REGION Network 28
   #temp := SCALE(IN := "5#净环热水阀门开度",
                  HI_LIM := 100.0,
                  LO_LIM := 0.0,
                  BIPOLAR := "AlwaysFALSE",
                  OUT => "AI"."5#净环热水阀门开度");
END_REGION

REGION Network 29
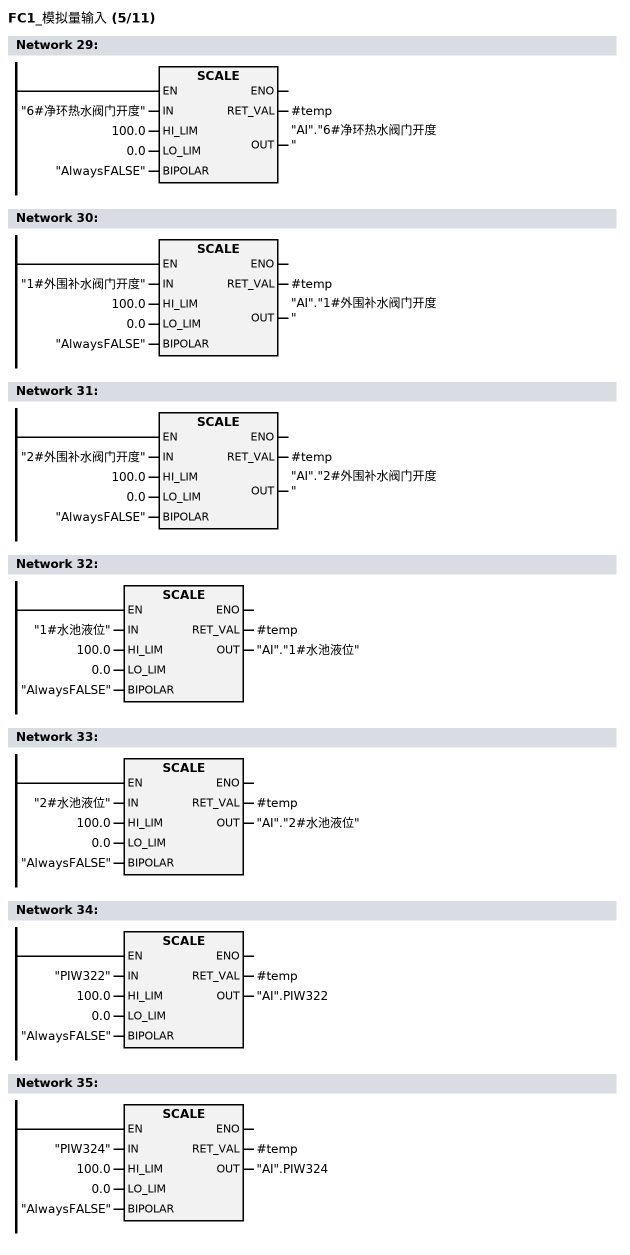
   #temp := SCALE(IN := "6#净环热水阀门开度",
                  HI_LIM := 100.0,
                  LO_LIM := 0.0,
                  BIPOLAR := "AlwaysFALSE",
                  OUT => "AI"."6#净环热水阀门开度");
END_REGION

REGION Network 30
   #temp := SCALE(IN := "1#外围补水阀门开度",
                  HI_LIM := 100.0,
                  LO_LIM := 0.0,
                  BIPOLAR := "AlwaysFALSE",
                  OUT => "AI"."1#外围补水阀门开度");
END_REGION

REGION Network 31
   #temp := SCALE(IN := "2#外围补水阀门开度",
                  HI_LIM := 100.0,
                  LO_LIM := 0.0,
                  BIPOLAR := "AlwaysFALSE",
                  OUT => "AI"."2#外围补水阀门开度");
END_REGION

REGION Network 32
   #temp := SCALE(IN := "1#水池液位",
                  HI_LIM := 100.0,
                  LO_LIM := 0.0,
                  BIPOLAR := "AlwaysFALSE",
                  OUT => "AI"."1#水池液位");
END_REGION

REGION Network 33
   #temp := SCALE(IN := "2#水池液位",
                  HI_LIM := 100.0,
                  LO_LIM := 0.0,
                  BIPOLAR := "AlwaysFALSE",
                  OUT => "AI"."2#水池液位");
END_REGION

REGION Network 34
   #temp := SCALE(IN := "PIW322", HI_LIM := 100.0, LO_LIM := 0.0, BIPOLAR := "AlwaysFALSE", OUT => "AI".PIW322);
END_REGION

REGION Network 35
   #temp := SCALE(IN := "PIW324", HI_LIM := 100.0, LO_LIM := 0.0, BIPOLAR := "AlwaysFALSE", OUT => "AI".PIW324);
END_REGION

REGION Network 36
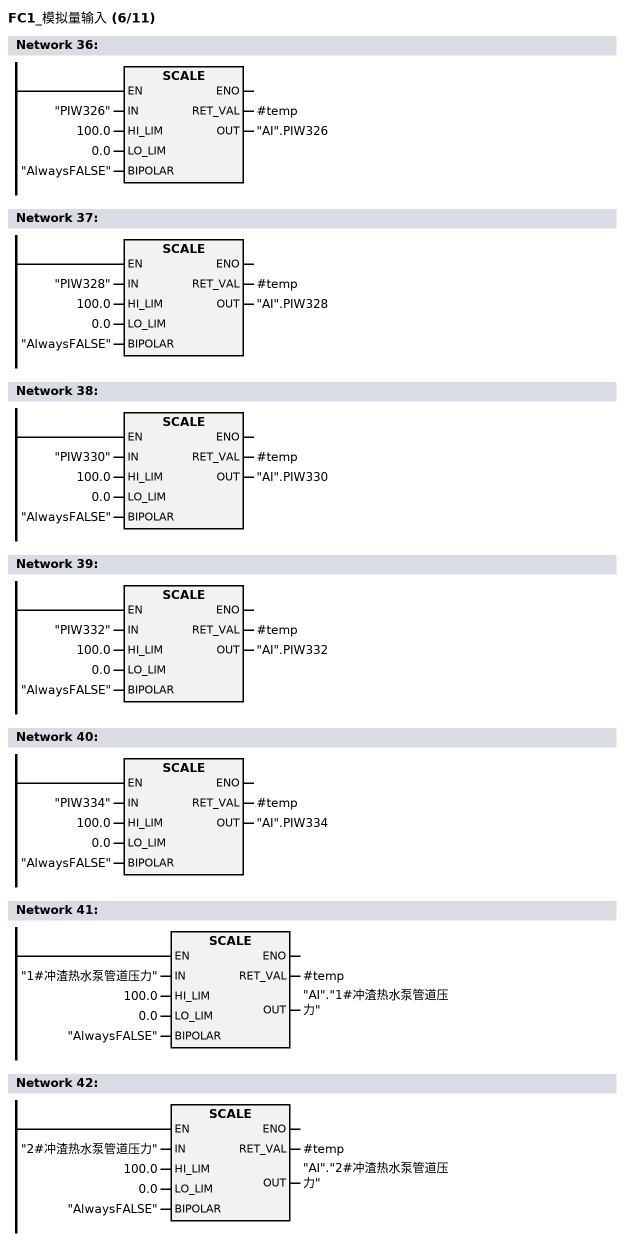
   #temp := SCALE(IN := "PIW326", HI_LIM := 100.0, LO_LIM := 0.0, BIPOLAR := "AlwaysFALSE", OUT => "AI".PIW326);
END_REGION

REGION Network 37
   #temp := SCALE(IN := "PIW328", HI_LIM := 100.0, LO_LIM := 0.0, BIPOLAR := "AlwaysFALSE", OUT => "AI".PIW328);
END_REGION

REGION Network 38
   #temp := SCALE(IN := "PIW330", HI_LIM := 100.0, LO_LIM := 0.0, BIPOLAR := "AlwaysFALSE", OUT => "AI".PIW330);
END_REGION

REGION Network 39
   #temp := SCALE(IN := "PIW332", HI_LIM := 100.0, LO_LIM := 0.0, BIPOLAR := "AlwaysFALSE", OUT => "AI".PIW332);
END_REGION

REGION Network 40
   #temp := SCALE(IN := "PIW334", HI_LIM := 100.0, LO_LIM := 0.0, BIPOLAR := "AlwaysFALSE", OUT => "AI".PIW334);
END_REGION

REGION Network 41
   #temp := SCALE(IN := "1#冲渣热水泵管道压力",
                  HI_LIM := 100.0,
                  LO_LIM := 0.0,
                  BIPOLAR := "AlwaysFALSE",
                  OUT => "AI"."1#冲渣热水泵管道压力");
END_REGION

REGION Network 42
   #temp := SCALE(IN := "2#冲渣热水泵管道压力",
                  HI_LIM := 100.0,
                  LO_LIM := 0.0,
                  BIPOLAR := "AlwaysFALSE",
                  OUT => "AI"."2#冲渣热水泵管道压力");
END_REGION

REGION Network 43
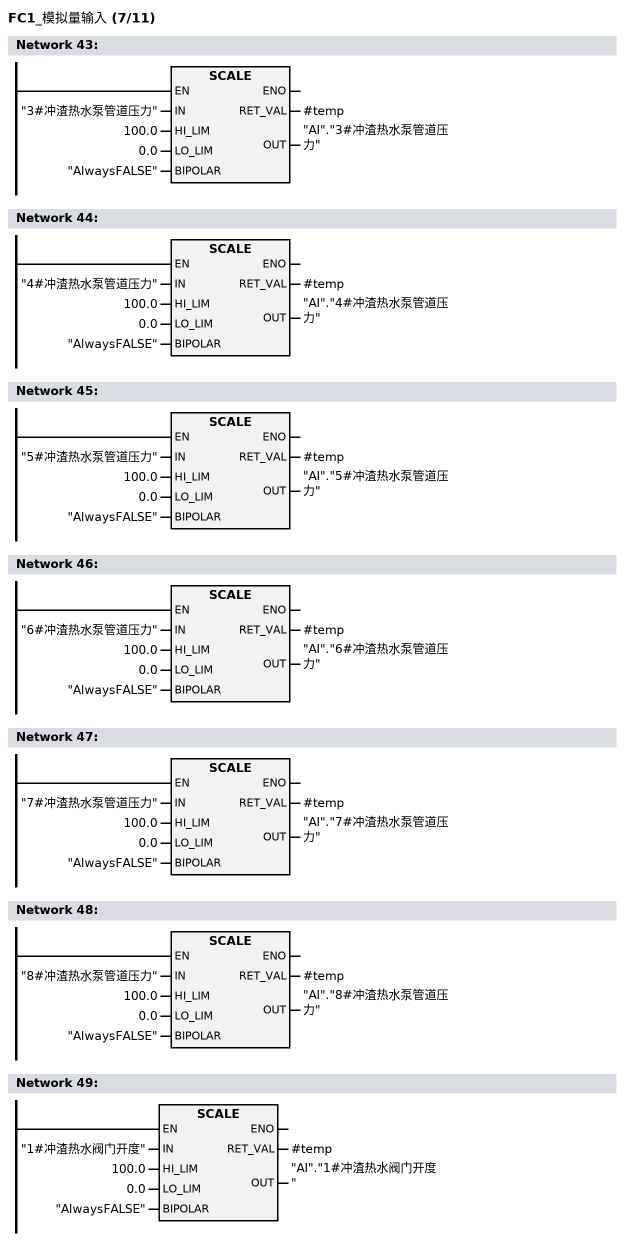
   #temp := SCALE(IN := "3#冲渣热水泵管道压力",
                  HI_LIM := 100.0,
                  LO_LIM := 0.0,
                  BIPOLAR := "AlwaysFALSE",
                  OUT => "AI"."3#冲渣热水泵管道压力");
END_REGION

REGION Network 44
   #temp := SCALE(IN := "4#冲渣热水泵管道压力",
                  HI_LIM := 100.0,
                  LO_LIM := 0.0,
                  BIPOLAR := "AlwaysFALSE",
                  OUT => "AI"."4#冲渣热水泵管道压力");
END_REGION

REGION Network 45
   #temp := SCALE(IN := "5#冲渣热水泵管道压力",
                  HI_LIM := 100.0,
                  LO_LIM := 0.0,
                  BIPOLAR := "AlwaysFALSE",
                  OUT => "AI"."5#冲渣热水泵管道压力");
END_REGION

REGION Network 46
   #temp := SCALE(IN := "6#冲渣热水泵管道压力",
                  HI_LIM := 100.0,
                  LO_LIM := 0.0,
                  BIPOLAR := "AlwaysFALSE",
                  OUT => "AI"."6#冲渣热水泵管道压力");
END_REGION

REGION Network 47
   #temp := SCALE(IN := "7#冲渣热水泵管道压力",
                  HI_LIM := 100.0,
                  LO_LIM := 0.0,
                  BIPOLAR := "AlwaysFALSE",
                  OUT => "AI"."7#冲渣热水泵管道压力");
END_REGION

REGION Network 48
   #temp := SCALE(IN := "8#冲渣热水泵管道压力",
                  HI_LIM := 100.0,
                  LO_LIM := 0.0,
                  BIPOLAR := "AlwaysFALSE",
                  OUT => "AI"."8#冲渣热水泵管道压力");
END_REGION

REGION Network 49
   #temp := SCALE(IN := "1#冲渣热水阀门开度",
                  HI_LIM := 100.0,
                  LO_LIM := 0.0,
                  BIPOLAR := "AlwaysFALSE",
                  OUT => "AI"."1#冲渣热水阀门开度");
END_REGION

REGION Network 50
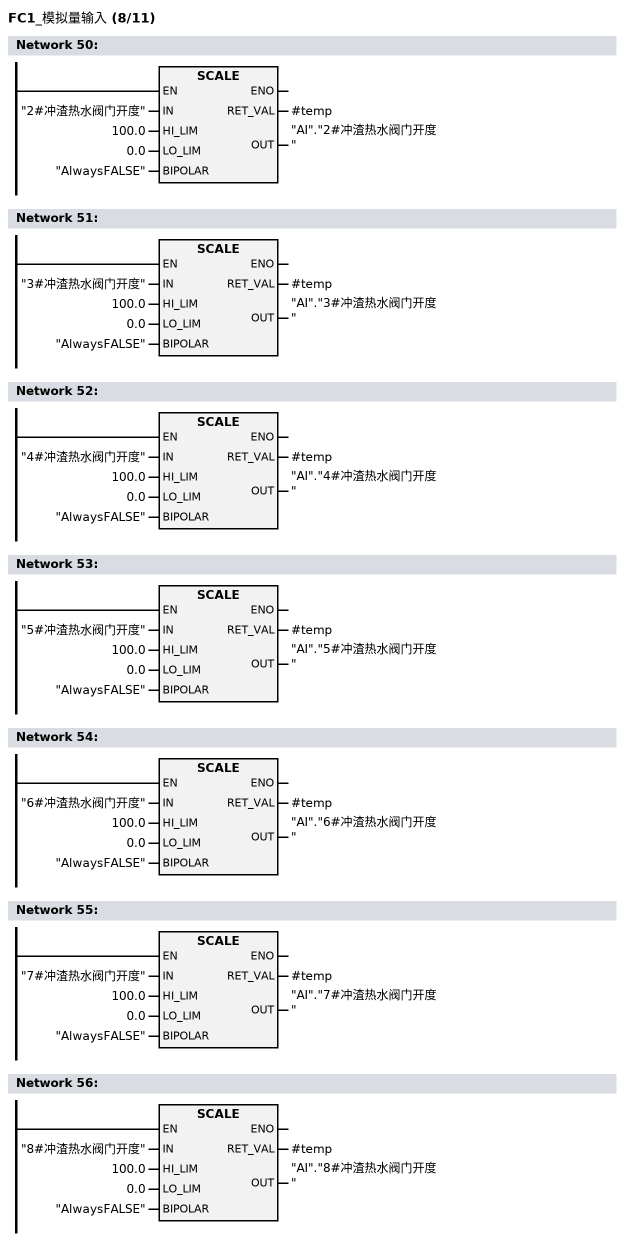
   #temp := SCALE(IN := "2#冲渣热水阀门开度",
                  HI_LIM := 100.0,
                  LO_LIM := 0.0,
                  BIPOLAR := "AlwaysFALSE",
                  OUT => "AI"."2#冲渣热水阀门开度");
END_REGION

REGION Network 51
   #temp := SCALE(IN := "3#冲渣热水阀门开度",
                  HI_LIM := 100.0,
                  LO_LIM := 0.0,
                  BIPOLAR := "AlwaysFALSE",
                  OUT => "AI"."3#冲渣热水阀门开度");
END_REGION

REGION Network 52
   #temp := SCALE(IN := "4#冲渣热水阀门开度",
                  HI_LIM := 100.0,
                  LO_LIM := 0.0,
                  BIPOLAR := "AlwaysFALSE",
                  OUT => "AI"."4#冲渣热水阀门开度");
END_REGION

REGION Network 53
   #temp := SCALE(IN := "5#冲渣热水阀门开度",
                  HI_LIM := 100.0,
                  LO_LIM := 0.0,
                  BIPOLAR := "AlwaysFALSE",
                  OUT => "AI"."5#冲渣热水阀门开度");
END_REGION

REGION Network 54
   #temp := SCALE(IN := "6#冲渣热水阀门开度",
                  HI_LIM := 100.0,
                  LO_LIM := 0.0,
                  BIPOLAR := "AlwaysFALSE",
                  OUT => "AI"."6#冲渣热水阀门开度");
END_REGION

REGION Network 55
   #temp := SCALE(IN := "7#冲渣热水阀门开度",
                  HI_LIM := 100.0,
                  LO_LIM := 0.0,
                  BIPOLAR := "AlwaysFALSE",
                  OUT => "AI"."7#冲渣热水阀门开度");
END_REGION

REGION Network 56
   #temp := SCALE(IN := "8#冲渣热水阀门开度",
                  HI_LIM := 100.0,
                  LO_LIM := 0.0,
                  BIPOLAR := "AlwaysFALSE",
                  OUT => "AI"."8#冲渣热水阀门开度");
END_REGION

REGION Network 57
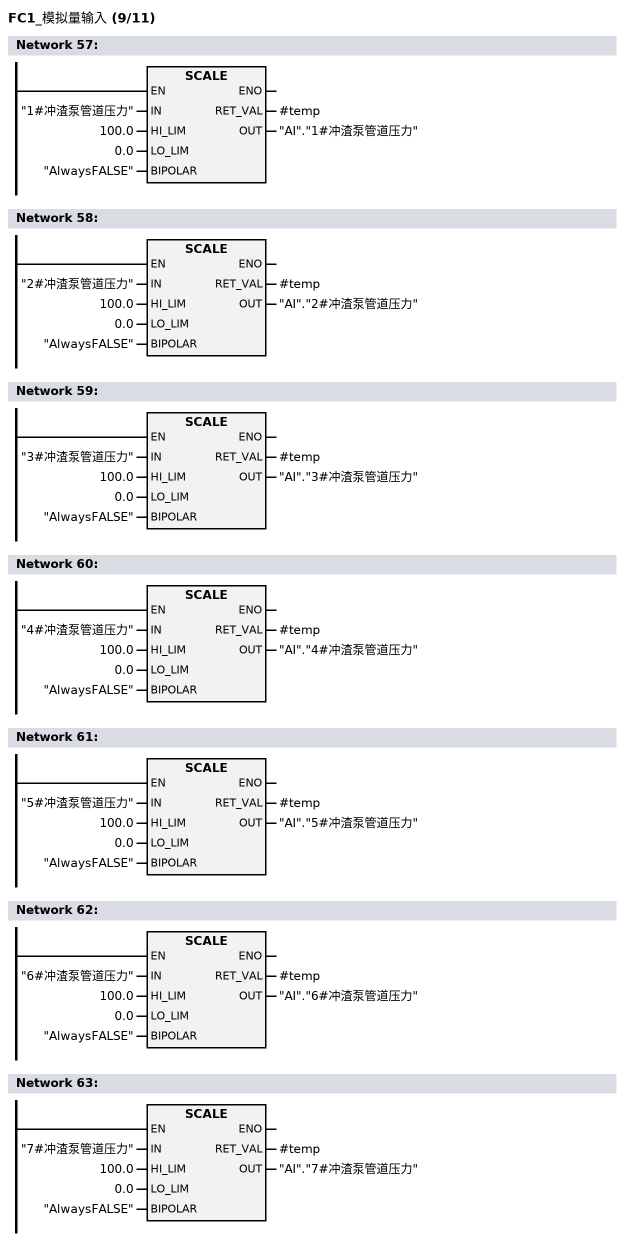
   #temp := SCALE(IN := "1#冲渣泵管道压力",
                  HI_LIM := 100.0,
                  LO_LIM := 0.0,
                  BIPOLAR := "AlwaysFALSE",
                  OUT => "AI"."1#冲渣泵管道压力");
END_REGION

REGION Network 58
   #temp := SCALE(IN := "2#冲渣泵管道压力",
                  HI_LIM := 100.0,
                  LO_LIM := 0.0,
                  BIPOLAR := "AlwaysFALSE",
                  OUT => "AI"."2#冲渣泵管道压力");
END_REGION

REGION Network 59
   #temp := SCALE(IN := "3#冲渣泵管道压力",
                  HI_LIM := 100.0,
                  LO_LIM := 0.0,
                  BIPOLAR := "AlwaysFALSE",
                  OUT => "AI"."3#冲渣泵管道压力");
END_REGION

REGION Network 60
   #temp := SCALE(IN := "4#冲渣泵管道压力",
                  HI_LIM := 100.0,
                  LO_LIM := 0.0,
                  BIPOLAR := "AlwaysFALSE",
                  OUT => "AI"."4#冲渣泵管道压力");
END_REGION

REGION Network 61
   #temp := SCALE(IN := "5#冲渣泵管道压力",
                  HI_LIM := 100.0,
                  LO_LIM := 0.0,
                  BIPOLAR := "AlwaysFALSE",
                  OUT => "AI"."5#冲渣泵管道压力");
END_REGION

REGION Network 62
   #temp := SCALE(IN := "6#冲渣泵管道压力",
                  HI_LIM := 100.0,
                  LO_LIM := 0.0,
                  BIPOLAR := "AlwaysFALSE",
                  OUT => "AI"."6#冲渣泵管道压力");
END_REGION

REGION Network 63
   #temp := SCALE(IN := "7#冲渣泵管道压力",
                  HI_LIM := 100.0,
                  LO_LIM := 0.0,
                  BIPOLAR := "AlwaysFALSE",
                  OUT => "AI"."7#冲渣泵管道压力");
END_REGION

REGION Network 64
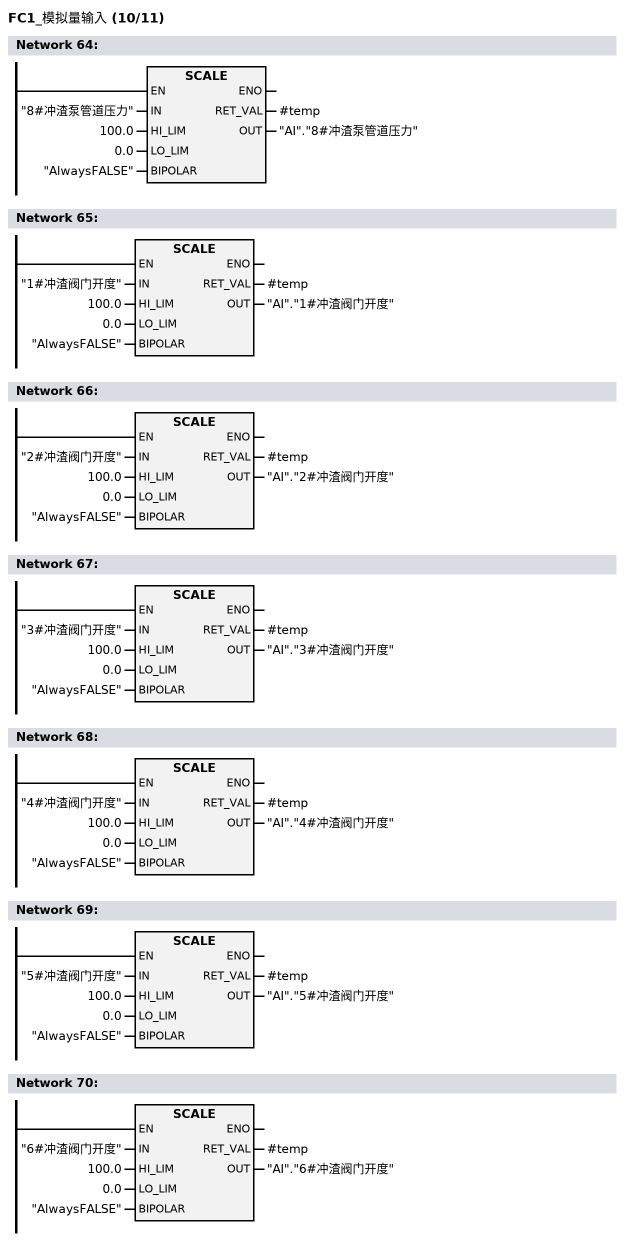
   #temp := SCALE(IN := "8#冲渣泵管道压力",
                  HI_LIM := 100.0,
                  LO_LIM := 0.0,
                  BIPOLAR := "AlwaysFALSE",
                  OUT => "AI"."8#冲渣泵管道压力");
END_REGION

REGION Network 65
   #temp := SCALE(IN := "1#冲渣阀门开度",
                  HI_LIM := 100.0,
                  LO_LIM := 0.0,
                  BIPOLAR := "AlwaysFALSE",
                  OUT => "AI"."1#冲渣阀门开度");
END_REGION

REGION Network 66
   #temp := SCALE(IN := "2#冲渣阀门开度",
                  HI_LIM := 100.0,
                  LO_LIM := 0.0,
                  BIPOLAR := "AlwaysFALSE",
                  OUT => "AI"."2#冲渣阀门开度");
END_REGION

REGION Network 67
   #temp := SCALE(IN := "3#冲渣阀门开度",
                  HI_LIM := 100.0,
                  LO_LIM := 0.0,
                  BIPOLAR := "AlwaysFALSE",
                  OUT => "AI"."3#冲渣阀门开度");
END_REGION

REGION Network 68
   #temp := SCALE(IN := "4#冲渣阀门开度",
                  HI_LIM := 100.0,
                  LO_LIM := 0.0,
                  BIPOLAR := "AlwaysFALSE",
                  OUT => "AI"."4#冲渣阀门开度");
END_REGION

REGION Network 69
   #temp := SCALE(IN := "5#冲渣阀门开度",
                  HI_LIM := 100.0,
                  LO_LIM := 0.0,
                  BIPOLAR := "AlwaysFALSE",
                  OUT => "AI"."5#冲渣阀门开度");
END_REGION

REGION Network 70
   #temp := SCALE(IN := "6#冲渣阀门开度",
                  HI_LIM := 100.0,
                  LO_LIM := 0.0,
                  BIPOLAR := "AlwaysFALSE",
                  OUT => "AI"."6#冲渣阀门开度");
END_REGION

REGION Network 71
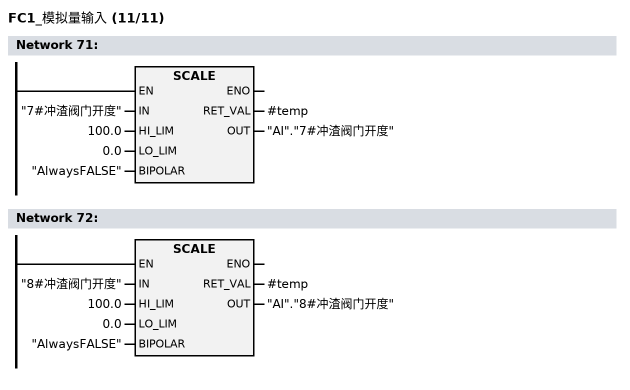
   #temp := SCALE(IN := "7#冲渣阀门开度",
                  HI_LIM := 100.0,
                  LO_LIM := 0.0,
                  BIPOLAR := "AlwaysFALSE",
                  OUT => "AI"."7#冲渣阀门开度");
END_REGION

REGION Network 72
   #temp := SCALE(IN := "8#冲渣阀门开度",
                  HI_LIM := 100.0,
                  LO_LIM := 0.0,
                  BIPOLAR := "AlwaysFALSE",
                  OUT => "AI"."8#冲渣阀门开度");
END_REGION
END_FUNCTION

FUNCTION "FC2_模拟量输出" : Void   // FC2, LAD
{ S7_Optimized_Access := 'TRUE' }
VERSION : 0.1
   VAR_TEMP
      temp_AO : Word;
   END_VAR
BEGIN

REGION Network 1
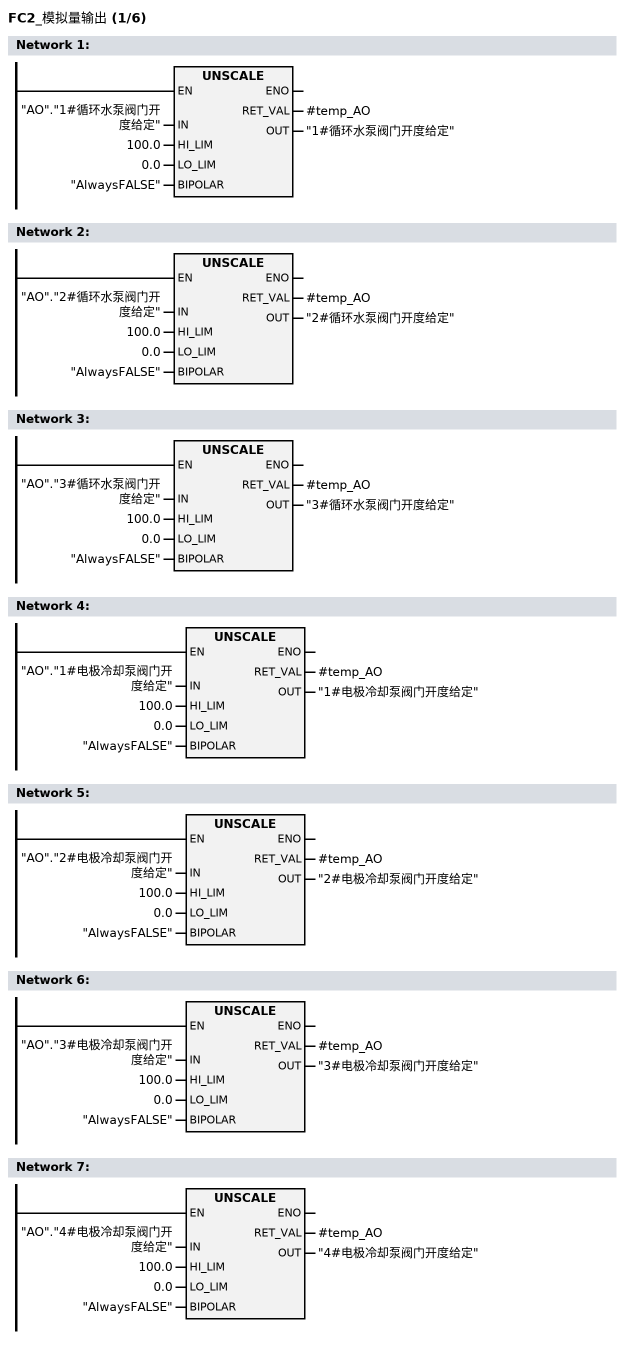
   #temp_AO := UNSCALE(IN := "AO"."1#循环水泵阀门开度给定",
                       HI_LIM := 100.0,
                       LO_LIM := 0.0,
                       BIPOLAR := "AlwaysFALSE",
                       OUT => "1#循环水泵阀门开度给定");
END_REGION

REGION Network 2
   #temp_AO := UNSCALE(IN := "AO"."2#循环水泵阀门开度给定",
                       HI_LIM := 100.0,
                       LO_LIM := 0.0,
                       BIPOLAR := "AlwaysFALSE",
                       OUT => "2#循环水泵阀门开度给定");
END_REGION

REGION Network 3
   #temp_AO := UNSCALE(IN := "AO"."3#循环水泵阀门开度给定",
                       HI_LIM := 100.0,
                       LO_LIM := 0.0,
                       BIPOLAR := "AlwaysFALSE",
                       OUT => "3#循环水泵阀门开度给定");
END_REGION

REGION Network 4
   #temp_AO := UNSCALE(IN := "AO"."1#电极冷却泵阀门开度给定",
                       HI_LIM := 100.0,
                       LO_LIM := 0.0,
                       BIPOLAR := "AlwaysFALSE",
                       OUT => "1#电极冷却泵阀门开度给定");
END_REGION

REGION Network 5
   #temp_AO := UNSCALE(IN := "AO"."2#电极冷却泵阀门开度给定",
                       HI_LIM := 100.0,
                       LO_LIM := 0.0,
                       BIPOLAR := "AlwaysFALSE",
                       OUT => "2#电极冷却泵阀门开度给定");
END_REGION

REGION Network 6
   #temp_AO := UNSCALE(IN := "AO"."3#电极冷却泵阀门开度给定",
                       HI_LIM := 100.0,
                       LO_LIM := 0.0,
                       BIPOLAR := "AlwaysFALSE",
                       OUT => "3#电极冷却泵阀门开度给定");
END_REGION

REGION Network 7
   #temp_AO := UNSCALE(IN := "AO"."4#电极冷却泵阀门开度给定",
                       HI_LIM := 100.0,
                       LO_LIM := 0.0,
                       BIPOLAR := "AlwaysFALSE",
                       OUT => "4#电极冷却泵阀门开度给定");
END_REGION

REGION Network 8
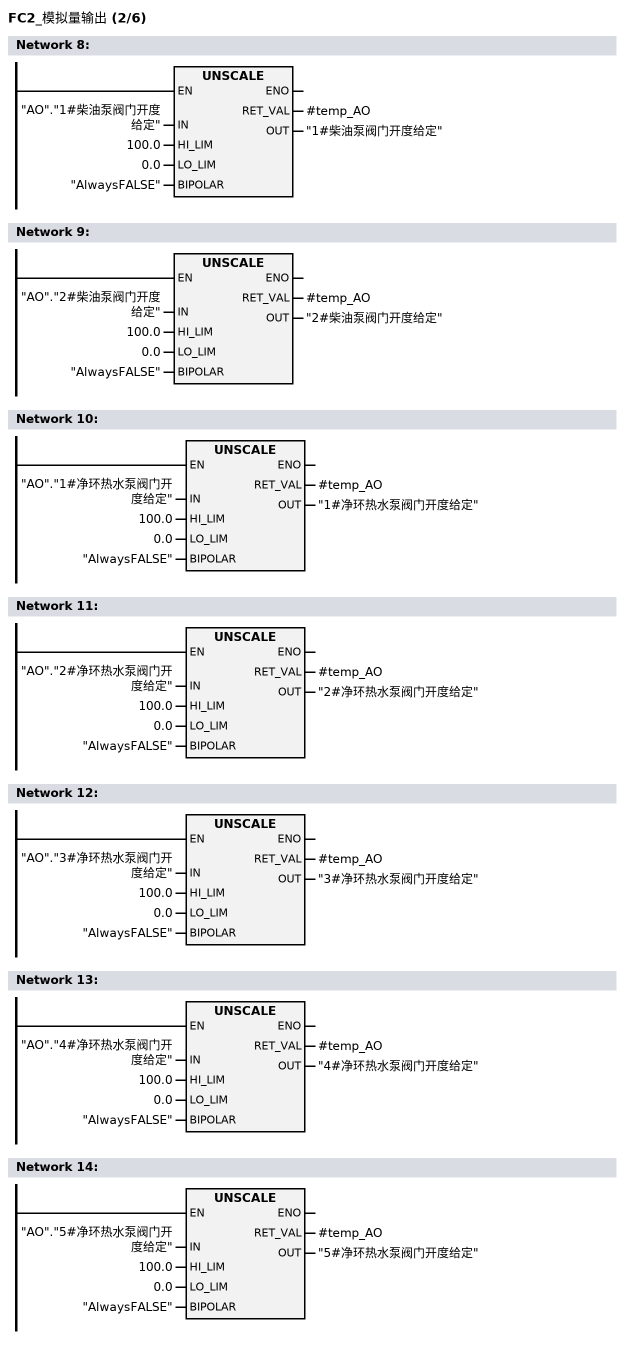
   #temp_AO := UNSCALE(IN := "AO"."1#柴油泵阀门开度给定",
                       HI_LIM := 100.0,
                       LO_LIM := 0.0,
                       BIPOLAR := "AlwaysFALSE",
                       OUT => "1#柴油泵阀门开度给定");
END_REGION

REGION Network 9
   #temp_AO := UNSCALE(IN := "AO"."2#柴油泵阀门开度给定",
                       HI_LIM := 100.0,
                       LO_LIM := 0.0,
                       BIPOLAR := "AlwaysFALSE",
                       OUT => "2#柴油泵阀门开度给定");
END_REGION

REGION Network 10
   #temp_AO := UNSCALE(IN := "AO"."1#净环热水泵阀门开度给定",
                       HI_LIM := 100.0,
                       LO_LIM := 0.0,
                       BIPOLAR := "AlwaysFALSE",
                       OUT => "1#净环热水泵阀门开度给定");
END_REGION

REGION Network 11
   #temp_AO := UNSCALE(IN := "AO"."2#净环热水泵阀门开度给定",
                       HI_LIM := 100.0,
                       LO_LIM := 0.0,
                       BIPOLAR := "AlwaysFALSE",
                       OUT => "2#净环热水泵阀门开度给定");
END_REGION

REGION Network 12
   #temp_AO := UNSCALE(IN := "AO"."3#净环热水泵阀门开度给定",
                       HI_LIM := 100.0,
                       LO_LIM := 0.0,
                       BIPOLAR := "AlwaysFALSE",
                       OUT => "3#净环热水泵阀门开度给定");
END_REGION

REGION Network 13
   #temp_AO := UNSCALE(IN := "AO"."4#净环热水泵阀门开度给定",
                       HI_LIM := 100.0,
                       LO_LIM := 0.0,
                       BIPOLAR := "AlwaysFALSE",
                       OUT => "4#净环热水泵阀门开度给定");
END_REGION

REGION Network 14
   #temp_AO := UNSCALE(IN := "AO"."5#净环热水泵阀门开度给定",
                       HI_LIM := 100.0,
                       LO_LIM := 0.0,
                       BIPOLAR := "AlwaysFALSE",
                       OUT => "5#净环热水泵阀门开度给定");
END_REGION

REGION Network 15
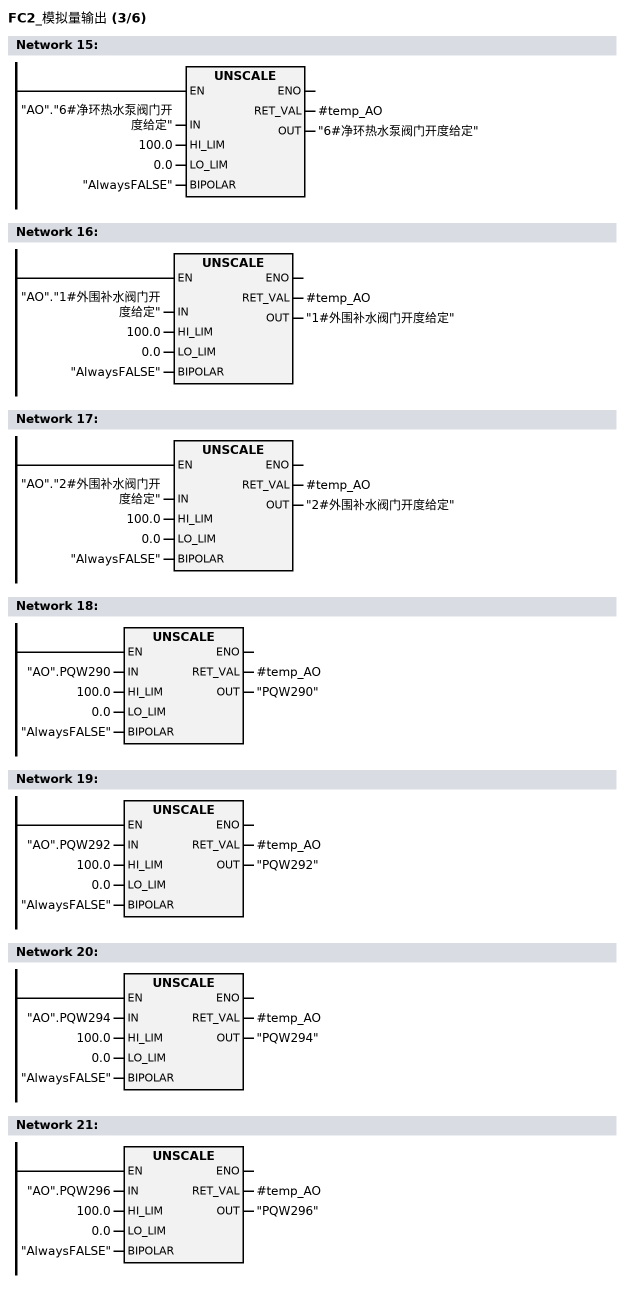
   #temp_AO := UNSCALE(IN := "AO"."6#净环热水泵阀门开度给定",
                       HI_LIM := 100.0,
                       LO_LIM := 0.0,
                       BIPOLAR := "AlwaysFALSE",
                       OUT => "6#净环热水泵阀门开度给定");
END_REGION

REGION Network 16
   #temp_AO := UNSCALE(IN := "AO"."1#外围补水阀门开度给定",
                       HI_LIM := 100.0,
                       LO_LIM := 0.0,
                       BIPOLAR := "AlwaysFALSE",
                       OUT => "1#外围补水阀门开度给定");
END_REGION

REGION Network 17
   #temp_AO := UNSCALE(IN := "AO"."2#外围补水阀门开度给定",
                       HI_LIM := 100.0,
                       LO_LIM := 0.0,
                       BIPOLAR := "AlwaysFALSE",
                       OUT => "2#外围补水阀门开度给定");
END_REGION

REGION Network 18
   #temp_AO := UNSCALE(IN := "AO".PQW290,
                       HI_LIM := 100.0,
                       LO_LIM := 0.0,
                       BIPOLAR := "AlwaysFALSE",
                       OUT => "PQW290");
END_REGION

REGION Network 19
   #temp_AO := UNSCALE(IN := "AO".PQW292,
                       HI_LIM := 100.0,
                       LO_LIM := 0.0,
                       BIPOLAR := "AlwaysFALSE",
                       OUT => "PQW292");
END_REGION

REGION Network 20
   #temp_AO := UNSCALE(IN := "AO".PQW294,
                       HI_LIM := 100.0,
                       LO_LIM := 0.0,
                       BIPOLAR := "AlwaysFALSE",
                       OUT => "PQW294");
END_REGION

REGION Network 21
   #temp_AO := UNSCALE(IN := "AO".PQW296,
                       HI_LIM := 100.0,
                       LO_LIM := 0.0,
                       BIPOLAR := "AlwaysFALSE",
                       OUT => "PQW296");
END_REGION

REGION Network 22
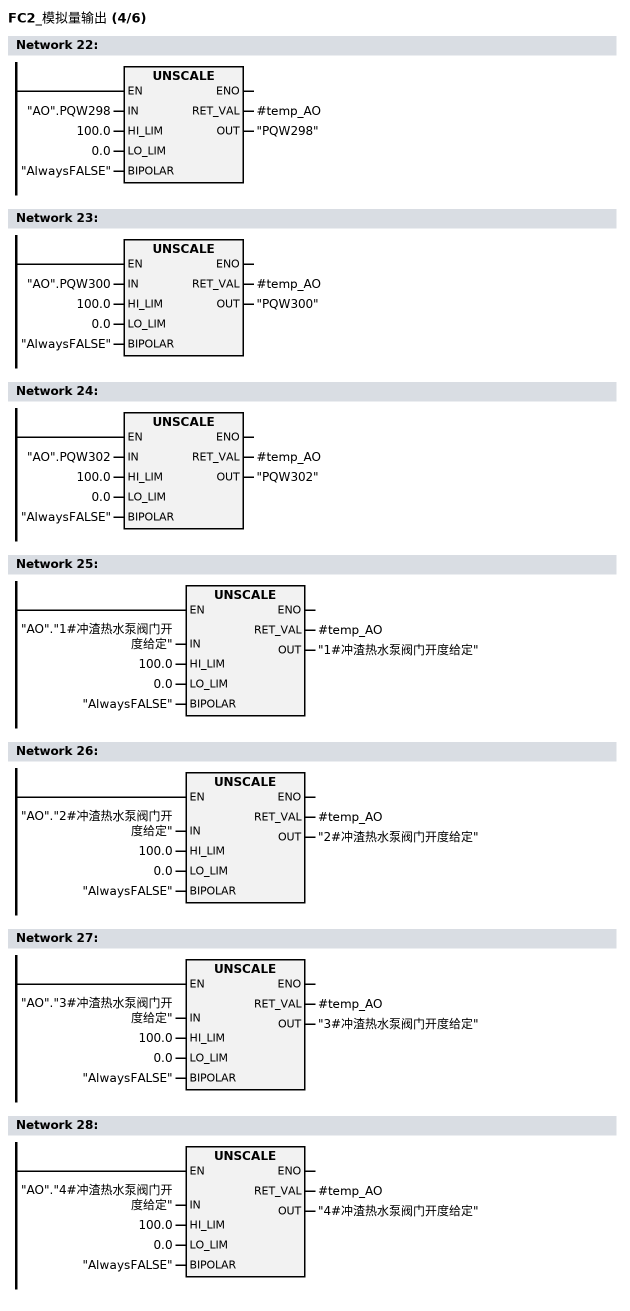
   #temp_AO := UNSCALE(IN := "AO".PQW298,
                       HI_LIM := 100.0,
                       LO_LIM := 0.0,
                       BIPOLAR := "AlwaysFALSE",
                       OUT => "PQW298");
END_REGION

REGION Network 23
   #temp_AO := UNSCALE(IN := "AO".PQW300,
                       HI_LIM := 100.0,
                       LO_LIM := 0.0,
                       BIPOLAR := "AlwaysFALSE",
                       OUT => "PQW300");
END_REGION

REGION Network 24
   #temp_AO := UNSCALE(IN := "AO".PQW302,
                       HI_LIM := 100.0,
                       LO_LIM := 0.0,
                       BIPOLAR := "AlwaysFALSE",
                       OUT => "PQW302");
END_REGION

REGION Network 25
   #temp_AO := UNSCALE(IN := "AO"."1#冲渣热水泵阀门开度给定",
                       HI_LIM := 100.0,
                       LO_LIM := 0.0,
                       BIPOLAR := "AlwaysFALSE",
                       OUT => "1#冲渣热水泵阀门开度给定");
END_REGION

REGION Network 26
   #temp_AO := UNSCALE(IN := "AO"."2#冲渣热水泵阀门开度给定",
                       HI_LIM := 100.0,
                       LO_LIM := 0.0,
                       BIPOLAR := "AlwaysFALSE",
                       OUT => "2#冲渣热水泵阀门开度给定");
END_REGION

REGION Network 27
   #temp_AO := UNSCALE(IN := "AO"."3#冲渣热水泵阀门开度给定",
                       HI_LIM := 100.0,
                       LO_LIM := 0.0,
                       BIPOLAR := "AlwaysFALSE",
                       OUT => "3#冲渣热水泵阀门开度给定");
END_REGION

REGION Network 28
   #temp_AO := UNSCALE(IN := "AO"."4#冲渣热水泵阀门开度给定",
                       HI_LIM := 100.0,
                       LO_LIM := 0.0,
                       BIPOLAR := "AlwaysFALSE",
                       OUT => "4#冲渣热水泵阀门开度给定");
END_REGION

REGION Network 29
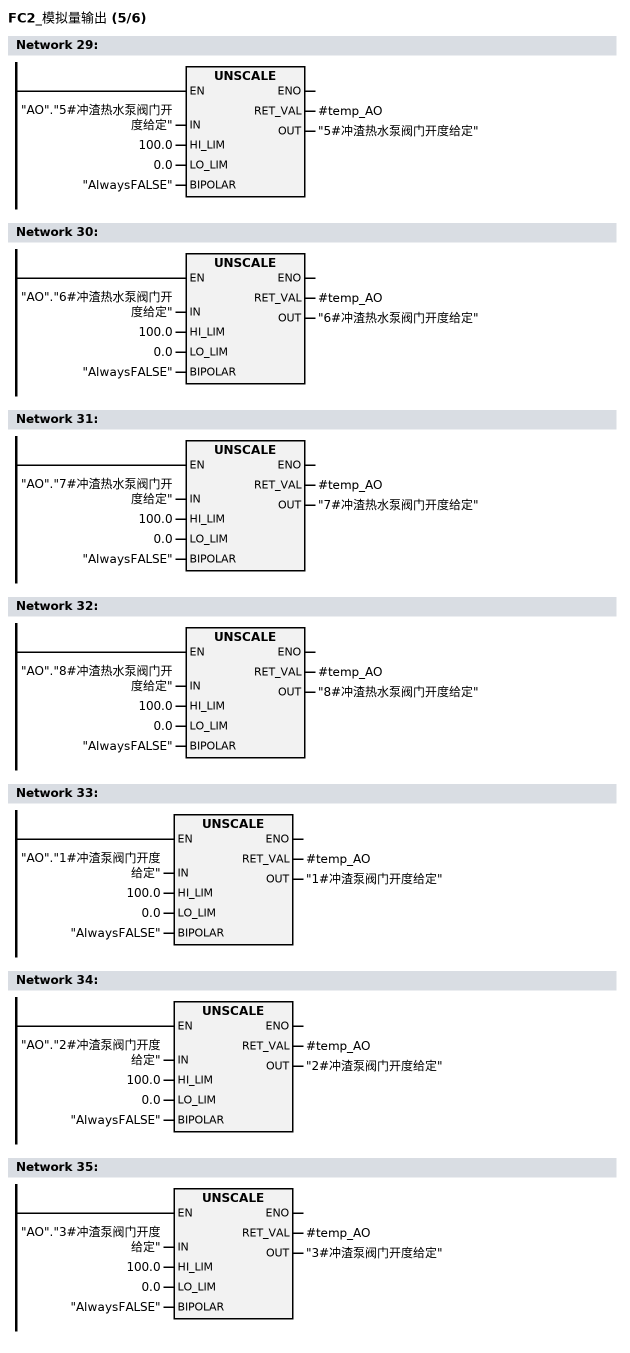
   #temp_AO := UNSCALE(IN := "AO"."5#冲渣热水泵阀门开度给定",
                       HI_LIM := 100.0,
                       LO_LIM := 0.0,
                       BIPOLAR := "AlwaysFALSE",
                       OUT => "5#冲渣热水泵阀门开度给定");
END_REGION

REGION Network 30
   #temp_AO := UNSCALE(IN := "AO"."6#冲渣热水泵阀门开度给定",
                       HI_LIM := 100.0,
                       LO_LIM := 0.0,
                       BIPOLAR := "AlwaysFALSE",
                       OUT => "6#冲渣热水泵阀门开度给定");
END_REGION

REGION Network 31
   #temp_AO := UNSCALE(IN := "AO"."7#冲渣热水泵阀门开度给定",
                       HI_LIM := 100.0,
                       LO_LIM := 0.0,
                       BIPOLAR := "AlwaysFALSE",
                       OUT => "7#冲渣热水泵阀门开度给定");
END_REGION

REGION Network 32
   #temp_AO := UNSCALE(IN := "AO"."8#冲渣热水泵阀门开度给定",
                       HI_LIM := 100.0,
                       LO_LIM := 0.0,
                       BIPOLAR := "AlwaysFALSE",
                       OUT => "8#冲渣热水泵阀门开度给定");
END_REGION

REGION Network 33
   #temp_AO := UNSCALE(IN := "AO"."1#冲渣泵阀门开度给定",
                       HI_LIM := 100.0,
                       LO_LIM := 0.0,
                       BIPOLAR := "AlwaysFALSE",
                       OUT => "1#冲渣泵阀门开度给定");
END_REGION

REGION Network 34
   #temp_AO := UNSCALE(IN := "AO"."2#冲渣泵阀门开度给定",
                       HI_LIM := 100.0,
                       LO_LIM := 0.0,
                       BIPOLAR := "AlwaysFALSE",
                       OUT => "2#冲渣泵阀门开度给定");
END_REGION

REGION Network 35
   #temp_AO := UNSCALE(IN := "AO"."3#冲渣泵阀门开度给定",
                       HI_LIM := 100.0,
                       LO_LIM := 0.0,
                       BIPOLAR := "AlwaysFALSE",
                       OUT => "3#冲渣泵阀门开度给定");
END_REGION

REGION Network 36
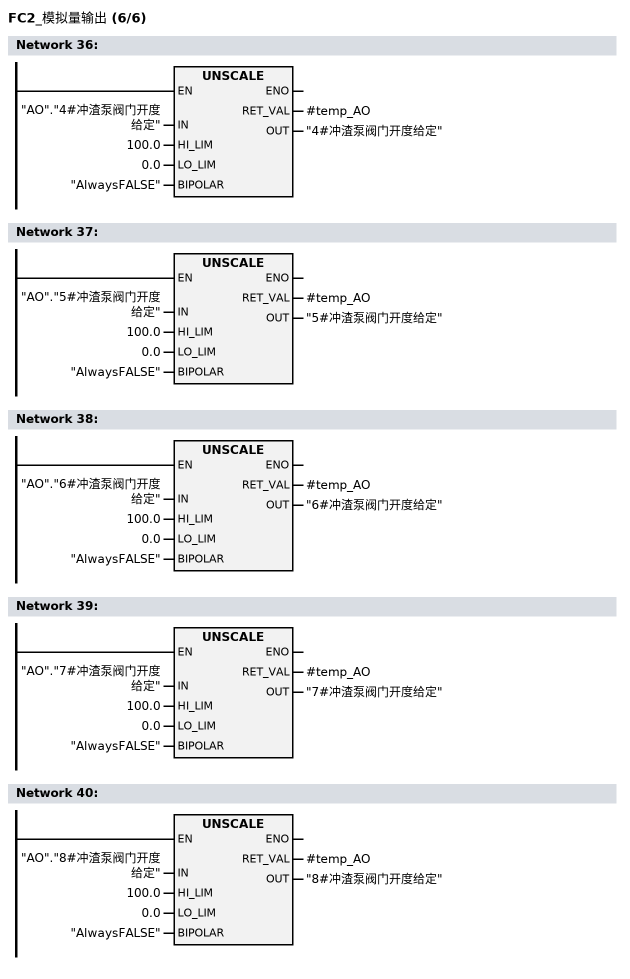
   #temp_AO := UNSCALE(IN := "AO"."4#冲渣泵阀门开度给定",
                       HI_LIM := 100.0,
                       LO_LIM := 0.0,
                       BIPOLAR := "AlwaysFALSE",
                       OUT => "4#冲渣泵阀门开度给定");
END_REGION

REGION Network 37
   #temp_AO := UNSCALE(IN := "AO"."5#冲渣泵阀门开度给定",
                       HI_LIM := 100.0,
                       LO_LIM := 0.0,
                       BIPOLAR := "AlwaysFALSE",
                       OUT => "5#冲渣泵阀门开度给定");
END_REGION

REGION Network 38
   #temp_AO := UNSCALE(IN := "AO"."6#冲渣泵阀门开度给定",
                       HI_LIM := 100.0,
                       LO_LIM := 0.0,
                       BIPOLAR := "AlwaysFALSE",
                       OUT => "6#冲渣泵阀门开度给定");
END_REGION

REGION Network 39
   #temp_AO := UNSCALE(IN := "AO"."7#冲渣泵阀门开度给定",
                       HI_LIM := 100.0,
                       LO_LIM := 0.0,
                       BIPOLAR := "AlwaysFALSE",
                       OUT => "7#冲渣泵阀门开度给定");
END_REGION

REGION Network 40
   #temp_AO := UNSCALE(IN := "AO"."8#冲渣泵阀门开度给定",
                       HI_LIM := 100.0,
                       LO_LIM := 0.0,
                       BIPOLAR := "AlwaysFALSE",
                       OUT => "8#冲渣泵阀门开度给定");
END_REGION
END_FUNCTION

FUNCTION "FC10_电机_冷却塔风机FC" : Void   // FC10, LAD
{ S7_Optimized_Access := 'TRUE' }
VERSION : 0.1
BEGIN

REGION Network 1
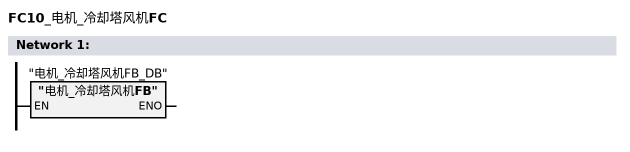
   RUNG wire#powerrail
      "电机_冷却塔风机FB_DB"()
   END_RUNG
   // the same network as SCL:
   "电机_冷却塔风机FB_DB"();   // "电机_冷却塔风机FB"
END_REGION
END_FUNCTION

FUNCTION "FC11_蝶阀FC" : Void   // FC11, LAD
{ S7_Optimized_Access := 'TRUE' }
VERSION : 0.1
BEGIN

REGION Network 1
